DATA_BLOCK "Library: Part Numbers as Text"   // DB3
{ S7_Optimized_Access := 'TRUE' }
VERSION : 0.1
BEGIN
   pnText[0] := WSTRING#'';
   pnText[1] := WSTRING#'11.52.001.0545.000B';
   pnText[2] := WSTRING#'11.52.001.315.000B';
   pnText[3] := WSTRING#'11.52.001.316.001D';
   pnText[4] := WSTRING#'11.54.007.045.015D';
   pnText[5] := WSTRING#'11.54.007.052.007B';
   pnText[6] := WSTRING#'11.54.007.052.008A';
   pnText[7] := WSTRING#'11.54.007.052.009B';
   pnText[8] := WSTRING#'11.54.007.052.010B';
   pnText[9] := WSTRING#'11.54.007.315.026G';
   pnText[10] := WSTRING#'11.54.017.315.001F';
   pnText[11] := WSTRING#'16.08.208.011.010G';
   pnText[12] := WSTRING#'16.08.208.021.020C';
   pnText[13] := WSTRING#'16.08.208.031.020C';
   pnText[14] := WSTRING#'16.08.208.041.000A';
   pnText[15] := WSTRING#'16.08.208.051.000A';
   pnText[16] := WSTRING#'16.08.208.081.010B';
   pnText[17] := WSTRING#'16.08.208.091.000A';
   pnText[18] := WSTRING#'16.08.208.101.010C';
   pnText[19] := WSTRING#'16.08.208.111.000B';
   pnText[20] := WSTRING#'16.08.208.131.010L';
   pnText[21] := WSTRING#'16.08.208.151.010F';
   pnText[22] := WSTRING#'16.08.208.161.020F';
   pnText[23] := WSTRING#'16.08.208.301.000F';
   pnText[24] := WSTRING#'16.08.208.311.000F';
   pnText[25] := WSTRING#'16.08.208.321.000G';
   pnText[26] := WSTRING#'16.08.208.331.000F';
   pnText[27] := WSTRING#'16.08.208.411.030C';
   pnText[28] := WSTRING#'16.08.208.501.000B';
   pnText[29] := WSTRING#'16.08.208.531.020L';
   pnText[30] := WSTRING#'16.08.208.621.010C';
   pnText[31] := WSTRING#'16.08.208.631.000F';
   pnText[32] := WSTRING#'16.08.208.651.010B';
   pnText[33] := WSTRING#'16.08.208.661.000F';
   pnText[34] := WSTRING#'16.08.208.691.010D';
   pnText[35] := WSTRING#'16.08.209.031.010C';
   pnText[36] := WSTRING#'16.08.209.031.030B';
   pnText[37] := WSTRING#'16.08.209.031.050A';
   pnText[38] := WSTRING#'16.08.209.091.010C';
   pnText[39] := WSTRING#'16.08.209.091.030D';
   pnText[40] := WSTRING#'16.08.209.091.060A';
   pnText[41] := WSTRING#'16.08.209.232.010C';
   pnText[42] := WSTRING#'16.08.210.031.010B';
   pnText[43] := WSTRING#'16.08.210.421.010A';
   pnText[44] := WSTRING#'16.08.210.421.020A';
   pnText[45] := WSTRING#'16.08.210.421.030A';
   pnText[46] := WSTRING#'16.08.211.121.000G';
   pnText[47] := WSTRING#'16.08.211.291.000A';
   pnText[48] := WSTRING#'16.08.211.511.020F';
   pnText[49] := WSTRING#'16.08.211.551.000B';
   pnText[50] := WSTRING#'16.08.211.781.000A';
   pnText[51] := WSTRING#'16.08.211.801.010A';
   pnText[52] := WSTRING#'16.08.211.801.020A';
   pnText[53] := WSTRING#'16.08.211.806.020A';
   pnText[54] := WSTRING#'16.08.215.141.010C';
   pnText[55] := WSTRING#'16.08.215.871.010C';
   pnText[56] := WSTRING#'16.08.216.011.030B';
   pnText[57] := WSTRING#'16.08.216.053.000A';
   pnText[58] := WSTRING#'16.08.216.057.001A';
   pnText[59] := WSTRING#'16.08.216.141.010C';
   pnText[60] := WSTRING#'16.08.216.151.010B';
   pnText[61] := WSTRING#'16.08.216.161.020A';
   pnText[62] := WSTRING#'16.08.216.181.010B';
   pnText[63] := WSTRING#'16.08.216.181.090A';
   pnText[64] := WSTRING#'16.08.216.181.100A';
   pnText[65] := WSTRING#'16.08.216.181.110B';
   pnText[66] := WSTRING#'16.08.216.200.050A';
   pnText[67] := WSTRING#'16.08.216.202.080A';
   pnText[68] := WSTRING#'16.08.216.231.000B';
   pnText[69] := WSTRING#'16.08.216.251.000B';
   pnText[70] := WSTRING#'16.08.216.291.000A';
   pnText[71] := WSTRING#'16.08.216.315.000A';
   pnText[72] := WSTRING#'16.08.216.315.001A';
   pnText[73] := WSTRING#'16.08.216.315.002A';
   pnText[74] := WSTRING#'16.08.216.501.000C';
   pnText[75] := WSTRING#'16.08.216.501.010A';
   pnText[76] := WSTRING#'16.08.216.511.000C';
   pnText[77] := WSTRING#'16.08.216.515.008C';
   pnText[78] := WSTRING#'16.08.216.521.000C';
   pnText[79] := WSTRING#'16.08.216.526.002C';
   pnText[80] := WSTRING#'16.08.216.526.009A';
   pnText[81] := WSTRING#'16.08.216.551.000B';
   pnText[82] := WSTRING#'16.08.216.722.001A';
   pnText[83] := WSTRING#'16.08.216.790.001A';
   pnText[84] := WSTRING#'16.08.216.806.020A';
   pnText[85] := WSTRING#'16.08.216.831.020A';
   pnText[86] := WSTRING#'16.08.216.871.010C';
   pnText[87] := WSTRING#'16.08.216.910.020B';
   pnText[88] := WSTRING#'16.08.216.911.000C';
   pnText[89] := WSTRING#'16.08.216.911.000G';
   pnText[90] := WSTRING#'16.08.216.911.000H';
   pnText[91] := WSTRING#'16.08.216.911.030B';
   pnText[92] := WSTRING#'16.08.216.911.040B';
   pnText[93] := WSTRING#'16.08.216.912.050A';
   pnText[94] := WSTRING#'16.08.216.912.060B';
   pnText[95] := WSTRING#'16.08.216.951.010A';
   pnText[96] := WSTRING#'16.08.216.181.020A';
   pnText[97] := WSTRING#'16.08.217.411.080A';
   pnText[98] := WSTRING#'16.08.217.421.010A';
   pnText[99] := WSTRING#'16.08.217.421.130A';
   pnText[100] := WSTRING#'16.18.007.301.010A';
   pnText[101] := WSTRING#'16.18.007.301.020A';
   pnText[102] := WSTRING#'16.18.007.311.010A';
   pnText[103] := WSTRING#'16.18.007.311.020A';
   pnText[104] := WSTRING#'16.18.007.321.010B';
   pnText[105] := WSTRING#'16.18.008.301.010A';
   pnText[106] := WSTRING#'16.18.008.301.020A';
   pnText[107] := WSTRING#'16.18.008.301.030A';
   pnText[108] := WSTRING#'16.18.008.311.010A';
   pnText[109] := WSTRING#'16.18.008.311.020B';
   pnText[110] := WSTRING#'16.18.009.301.010A';
   pnText[111] := WSTRING#'16.18.009.301.020B';
   pnText[112] := WSTRING#'16.18.009.301.030A';
   pnText[113] := WSTRING#'16.18.009.301.040B';
   pnText[114] := WSTRING#'16.18.009.301.050A';
   pnText[115] := WSTRING#'16.18.009.311.010A';
   pnText[116] := WSTRING#'16.18.009.321.010A';
   pnText[117] := WSTRING#'16.18.009.321.020B';
   pnText[118] := WSTRING#'16.18.009.321.030A';
   pnText[119] := WSTRING#'16.18.009.331.030A';
   pnText[120] := WSTRING#'16.18.009.331.050A';
   pnText[121] := WSTRING#'16.18.009.371.010A';
   pnText[122] := WSTRING#'16.18.011.301.010A';
   pnText[123] := WSTRING#'16.18.011.301.020B';
   pnText[124] := WSTRING#'16.18.011.301.030A';
   pnText[125] := WSTRING#'16.18.011.301.040B';
   pnText[126] := WSTRING#'16.18.011.311.020A';
   pnText[127] := WSTRING#'16.18.011.321.010A';
   pnText[128] := WSTRING#'16.18.011.321.020B';
   pnText[129] := WSTRING#'16.18.011.321.030A';
   pnText[130] := WSTRING#'16.18.011.331.010A';
   pnText[131] := WSTRING#'16.18.011.331.020D';
   pnText[132] := WSTRING#'16.18.012.401.010A';
   pnText[133] := WSTRING#'16.18.012.401.020A';
   pnText[134] := WSTRING#'16.18.012.411.010A';
   pnText[135] := WSTRING#'16.18.012.411.020B';
   pnText[136] := WSTRING#'16.18.012.431.010A';
   pnText[137] := WSTRING#'16.18.012.441.010A';
   pnText[138] := WSTRING#'16.18.013.411.010A';
   pnText[139] := WSTRING#'16.18.013.411.020B';
   pnText[140] := WSTRING#'16.18.013.411.030A';
   pnText[141] := WSTRING#'16.18.013.421.010A';
   pnText[142] := WSTRING#'16.18.014.411.010A';
   pnText[143] := WSTRING#'16.18.014.411.030A';
   pnText[144] := WSTRING#'16.18.015.401.010A';
   pnText[145] := WSTRING#'16.18.015.411.010A';
   pnText[146] := WSTRING#'16.18.015.411.020B';
   pnText[147] := WSTRING#'16.18.015.411.030A';
   pnText[148] := WSTRING#'16.18.015.421.010A';
   pnText[149] := WSTRING#'16.18.015.421.020B';
   pnText[150] := WSTRING#'16.18.017.301.010A';
   pnText[151] := WSTRING#'16.18.017.301.020A';
   pnText[152] := WSTRING#'16.18.017.301.030A';
   pnText[153] := WSTRING#'16.18.017.301.040A';
   pnText[154] := WSTRING#'16.18.017.301.050A';
   pnText[155] := WSTRING#'16.18.017.311.010A';
   pnText[156] := WSTRING#'16.18.017.321.010A';
   pnText[157] := WSTRING#'16.18.017.321.020A';
   pnText[158] := WSTRING#'16.18.018.400.000A';
   pnText[159] := WSTRING#'16.18.018.401.010A';
   pnText[160] := WSTRING#'16.18.018.401.020B';
   pnText[161] := WSTRING#'16.18.018.401.030A';
   pnText[162] := WSTRING#'16.18.018.411.010A';
   pnText[163] := WSTRING#'16.18.018.421.010B';
   pnText[164] := WSTRING#'16.32.112.054.041A';
   pnText[165] := WSTRING#'16.32.112.057.010A';
   pnText[166] := WSTRING#'16.32.112.500.060D';
   pnText[167] := WSTRING#'16.32.112.500.090B';
   pnText[168] := WSTRING#'16.32.112.500.100A';
   pnText[169] := WSTRING#'16.32.112.500.120A';
   pnText[170] := WSTRING#'16.32.112.500.150B';
   pnText[171] := WSTRING#'16.32.112.500.160A';
   pnText[172] := WSTRING#'16.32.112.500.220A';
   pnText[173] := WSTRING#'16.32.112.500.300E';
   pnText[174] := WSTRING#'16.32.112.500.520B';
   pnText[175] := WSTRING#'16.32.112.502.050B';
   pnText[176] := WSTRING#'16.32.112.502.060B';
   pnText[177] := WSTRING#'16.32.112.502.070E';
   pnText[178] := WSTRING#'16.32.112.503.210A';
   pnText[179] := WSTRING#'16.32.112.503.220A';
   pnText[180] := WSTRING#'16.32.112.504.060A';
   pnText[181] := WSTRING#'16.32.112.504.070G';
   pnText[182] := WSTRING#'16.32.112.509.050E';
   pnText[183] := WSTRING#'16.32.112.509.070A';
   pnText[184] := WSTRING#'16.32.112.509.080F';
   pnText[185] := WSTRING#'16.32.112.516.110E';
   pnText[186] := WSTRING#'16.32.112.520.300E';
   pnText[187] := WSTRING#'16.32.112.521.010B';
   pnText[188] := WSTRING#'16.32.112.521.020B';
   pnText[189] := WSTRING#'16.32.112.521.030A';
   pnText[190] := WSTRING#'16.32.112.522.040D';
   pnText[191] := WSTRING#'16.32.112.522.050A';
   pnText[192] := WSTRING#'16.32.112.522.130A';
   pnText[193] := WSTRING#'16.32.112.529.010A';
   pnText[194] := WSTRING#'16.32.112.529.020B';
   pnText[195] := WSTRING#'16.32.112.529.030A';
   pnText[196] := WSTRING#'16.32.112.529.050D';
   pnText[197] := WSTRING#'16.32.112.536.010A';
   pnText[198] := WSTRING#'16.32.112.543.020A';
   pnText[199] := WSTRING#'16.32.112.543.210E';
   pnText[200] := WSTRING#'16.32.112.553.010A';
   pnText[201] := WSTRING#'16.32.112.553.020A';
   pnText[202] := WSTRING#'16.32.112.553.100D';
   pnText[203] := WSTRING#'16.32.112.553.220A';
   pnText[204] := WSTRING#'16.32.112.580.020A';
   pnText[205] := WSTRING#'16.32.112.601.030A';
   pnText[206] := WSTRING#'16.32.112.601.040A';
   pnText[207] := WSTRING#'16.32.112.621.010A';
   pnText[208] := WSTRING#'16.32.112.621.020A';
   pnText[209] := WSTRING#'16.32.112.704.000C';
   pnText[210] := WSTRING#'16.32.112.751.000D';
   pnText[211] := WSTRING#'16.32.112.751.001C';
   pnText[212] := WSTRING#'16.32.112.757.000A';
   pnText[213] := WSTRING#'16.32.112.757.001A';
   pnText[214] := WSTRING#'16.32.112.851.000A';
   pnText[215] := WSTRING#'16.32.112.851.001A';
   pnText[216] := WSTRING#'16.32.112.870.000C';
   pnText[217] := WSTRING#'16.32.307.211.150B';
   pnText[218] := WSTRING#'16.32.307.211.170B';
   pnText[219] := WSTRING#'16.32.307.212.320C';
   pnText[220] := WSTRING#'16.32.307.232.300B';
   pnText[221] := WSTRING#'16.32.307.262.300B';
   pnText[222] := WSTRING#'16.32.307.312.310A';
   pnText[223] := WSTRING#'16.32.307.461.160A';
   pnText[224] := WSTRING#'16.32.407.241.150B';
   pnText[225] := WSTRING#'16.32.407.241.170B';
   pnText[226] := WSTRING#'16.32.407.441.160A';
   pnText[227] := WSTRING#'16.32.606.311.010C';
   pnText[228] := WSTRING#'16.32.606.311.040B';
   pnText[229] := WSTRING#'16.32.606.311.050B';
   pnText[230] := WSTRING#'16.32.606.311.060A';
   pnText[231] := WSTRING#'16.32.606.311.070A';
   pnText[232] := WSTRING#'16.32.606.321.010B';
   pnText[233] := WSTRING#'16.32.606.321.030B';
   pnText[234] := WSTRING#'16.32.706.311.010C';
   pnText[235] := WSTRING#'16.32.706.311.020B';
   pnText[236] := WSTRING#'16.32.706.311.040B';
   pnText[237] := WSTRING#'16.32.706.311.050B';
   pnText[238] := WSTRING#'16.32.706.321.010B';
   pnText[239] := WSTRING#'16.32.706.321.030B';
   pnText[240] := WSTRING#'16.32.706.401.040A';
   pnText[241] := WSTRING#'16.32.706.401.050A';
   pnText[242] := WSTRING#'16.32.806.502.080A';
   pnText[243] := WSTRING#'DUNNAGE';
   pnText[244] := WSTRING#'PEANUTS';
   pnText[245] := WSTRING#'RINGS CART';
END_DATA_BLOCK

DATA_BLOCK "LED Sign"   // DB4
{ S7_Optimized_Access := 'TRUE' }
VERSION : 0.1
   VAR
      request : "LED Sign Data";
   END_VAR
BEGIN
END_DATA_BLOCK

DATA_BLOCK "HMI Stations: Saved Wips"   // DB5
{ S7_Optimized_Access := 'TRUE' }
VERSION : 0.1
BEGIN
   stn[0].pStn := 25;
   stn[1].pStn := 26;
   stn[2].pStn := 27;
   stn[3].pStn := 28;
   stn[4].pStn := 29;
END_DATA_BLOCK

DATA_BLOCK "HMI Data: TP700 Stations"   // DB6
{ S7_Optimized_Access := 'TRUE' }
VERSION : 0.1
BEGIN
END_DATA_BLOCK

DATA_BLOCK "Library: Wip Names as Text"   // DB8
{ S7_Optimized_Access := 'TRUE' }
VERSION : 0.1
BEGIN
   code[0] := WSTRING#'';
   code[1] := WSTRING#'11.52.001.312.000B';
   code[2] := WSTRING#'11.54.007.309.000D';
   code[3] := WSTRING#'11.54.007.309.002D';
   code[4] := WSTRING#'16.08.208.031.000F';
   code[5] := WSTRING#'16.08.208.081.000H';
   code[6] := WSTRING#'16.08.208.101.020A';
   code[7] := WSTRING#'16.08.208.621.000G';
   code[8] := WSTRING#'16.08.208.651.000G';
   code[9] := WSTRING#'16.08.209.031.000C';
   code[10] := WSTRING#'16.08.209.091.000D';
   code[11] := WSTRING#'16.08.209.233.000E';
   code[12] := WSTRING#'16.08.209.437.000A';
   code[13] := WSTRING#'16.08.210.031.000B';
   code[14] := WSTRING#'16.08.210.421.500A';
   code[15] := WSTRING#'16.08.210.428.000A';
   code[16] := WSTRING#'16.08.211.801.400A';
   code[17] := WSTRING#'16.08.211.801.700B';
   code[18] := WSTRING#'16.08.211.803.400A';
   code[19] := WSTRING#'16.08.211.806.400B';
   code[20] := WSTRING#'16.08.216.751.100A';
   code[21] := WSTRING#'16.08.216.801.600A';
   code[22] := WSTRING#'16.08.216.806.400A';
   code[23] := WSTRING#'16.08.217.233.000A';
   code[24] := WSTRING#'16.08.217.408.000A';
   code[25] := WSTRING#'16.08.217.421.500A';
   code[26] := WSTRING#'16.08.217.737.000A';
   code[27] := WSTRING#'16.18.007.300.000A';
   code[28] := WSTRING#'16.18.007.310.000A';
   code[29] := WSTRING#'16.18.007.320.000B';
   code[30] := WSTRING#'16.18.008.300.000A';
   code[31] := WSTRING#'16.18.008.310.000A';
   code[32] := WSTRING#'16.18.008.320.000A';
   code[33] := WSTRING#'16.18.008.340.000A';
   code[34] := WSTRING#'16.18.009.301.000H';
   code[35] := WSTRING#'16.18.009.311.000H';
   code[36] := WSTRING#'16.18.009.321.000G';
   code[37] := WSTRING#'16.18.009.331.000F';
   code[38] := WSTRING#'16.18.009.371.000D';
   code[39] := WSTRING#'16.18.011.300.000A';
   code[40] := WSTRING#'16.18.011.310.000A';
   code[41] := WSTRING#'16.18.011.320.000A';
   code[42] := WSTRING#'16.18.011.330.000A';
   code[43] := WSTRING#'16.18.011.340.000A';
   code[44] := WSTRING#'16.18.012.400.000A';
   code[45] := WSTRING#'16.18.012.410.000A';
   code[46] := WSTRING#'16.18.012.420.000A';
   code[47] := WSTRING#'16.18.012.430.000A';
   code[48] := WSTRING#'16.18.012.440.000A';
   code[49] := WSTRING#'16.18.013.410.000A';
   code[50] := WSTRING#'16.18.013.420.000A';
   code[51] := WSTRING#'16.18.015.400.000A';
   code[52] := WSTRING#'16.18.015.410.000A';
   code[53] := WSTRING#'16.18.015.420.000A';
   code[54] := WSTRING#'16.18.015.430.000A';
   code[55] := WSTRING#'16.18.015.450.000A';
   code[56] := WSTRING#'16.18.016.400.000A';
   code[57] := WSTRING#'16.18.017.300.000A';
   code[58] := WSTRING#'16.18.017.310.000A';
   code[59] := WSTRING#'16.18.017.321.000F';
   code[60] := WSTRING#'16.18.018.400.000A';
   code[61] := WSTRING#'16.18.018.410.000A';
   code[62] := WSTRING#'16.18.018.420.000A';
   code[63] := WSTRING#'16.18.018.440.000A';
   code[64] := WSTRING#'16.32.112.304.008A';
   code[65] := WSTRING#'16.32.112.311.001A';
   code[66] := WSTRING#'16.32.112.516.000G';
   code[67] := WSTRING#'16.32.112.543.000E';
   code[68] := WSTRING#'16.32.112.553.300C';
   code[69] := WSTRING#'16.32.307.322.210A';
   code[70] := WSTRING#'16.32.307.332.300A';
   code[71] := WSTRING#'16.32.307.332.400A';
   code[72] := WSTRING#'16.32.307.472.210A';
   code[73] := WSTRING#'16.32.407.322.210A';
   code[74] := WSTRING#'16.32.407.322.300A';
   code[75] := WSTRING#'16.32.606.411.000A';
   code[76] := WSTRING#'16.32.606.421.000A';
   code[77] := WSTRING#'16.32.706.311.000A';
   code[78] := WSTRING#'16.32.706.311.001A';
   code[79] := WSTRING#'16.32.706.341.000A';
   code[80] := WSTRING#'16.32.706.401.000A';
   txt[0] := WSTRING#'NO TEXT ENTERED';
   txt[1] := WSTRING#'DPF Sleeved 2016';
   txt[2] := WSTRING#'SA SCR CANNING 9.5 x 10in -END FORMED-';
   txt[3] := WSTRING#'Assembly DPF Canning 2016';
   txt[4] := WSTRING#'ASSY DOC CANNING A700';
   txt[5] := WSTRING#'ASSY DPF CANNING A700';
   txt[6] := WSTRING#'ASSY SCR CANNING FORMED';
   txt[7] := WSTRING#'DOC Stuffed Shell Before Forming';
   txt[8] := WSTRING#'DOC Stuffed Shell Unformed';
   txt[9] := WSTRING#'DPF Stuffed Shell 1 box longs only';
   txt[10] := WSTRING#'DPF Stuffed Shell MD11';
   txt[11] := WSTRING#'DPF Stuffed Shell: MD13/MD16';
   txt[12] := WSTRING#'SA DOC CANNING 11.25 x 3.4in -END FORMED';
   txt[13] := WSTRING#'SA DOC CANNING 11.25 x 4in -END FORMED-';
   txt[14] := WSTRING#'SA DOC CANNING 11.25 x 5in -END FORMED-';
   txt[15] := WSTRING#'SA DOC CANNING 11.25 x 6.8in -END FORMED';
   txt[16] := WSTRING#'SA DOC CANNING 11_25 x 5in -END FORMED-';
   txt[17] := WSTRING#'SA DOC CANNING 9.5 x 3.3in -END FORMED-';
   txt[18] := WSTRING#'SA DOC CANNING 9.5 x 4in -END FORMED-';
   txt[19] := WSTRING#'SA DOC CANNING 9.5 x 4in -END FORMED_';
   txt[20] := WSTRING#'SA DOC CANNING 9.5 x 5.5in -END FORMED-';
   txt[21] := WSTRING#'SA DOC CANNING 9.5 x 5in -END FORMED-';
   txt[22] := WSTRING#'SA DOC CANNING 9_5 x 4_5in -END FORMED-';
   txt[23] := WSTRING#'SA DOC Canning w/out End Forming';
   txt[24] := WSTRING#'SA DOC Sleeved';
   txt[25] := WSTRING#'SA DOC SLEEVED - 2HH 2016';
   txt[26] := WSTRING#'SA DOC SLEEVED - 2V2 2016 unformed';
   txt[27] := WSTRING#'SA DOC Sleeved Before Forming';
   txt[28] := WSTRING#'SA DOC Sleeved DDC 2016 unformed';
   txt[29] := WSTRING#'SA DPF SLEEVED Hess';
   txt[30] := WSTRING#'SA DPF Stuffed (after Hess)';
   txt[31] := WSTRING#'SA DPF Stuffed Shell';
   txt[32] := WSTRING#'SA JL 2.2L DPF CANNING';
   txt[33] := WSTRING#'SA SCR CANNING 12 x 10in -END FORMED-';
   txt[34] := WSTRING#'SA SCR CANNING 12 x 9in -END FORMED-';
   txt[35] := WSTRING#'SA SCR CANNING 12x7in UNFORMED-';
   txt[36] := WSTRING#'SA SCR CANNING 13 x 11in UNFORMED-';
   txt[37] := WSTRING#'SA SCR CANNING 13 x 12in UNFORMED-';
   txt[38] := WSTRING#'SA SCR CANNING 13 x 9in UNFORMED';
   txt[39] := WSTRING#'SA SCR CANNING 13 X10 UNFORMED';
   txt[40] := WSTRING#'SA SCR CANNING 9.5 x 10in -END FORMED-';
   txt[41] := WSTRING#'SA SCR CANNING 9.5 x 12in -END FORMED-';
   txt[42] := WSTRING#'SA SCR CANNING 9.5 x 13.5in -END FORMED-';
   txt[43] := WSTRING#'SA SCR CANNING 9.5 x 13in -END FORMED-';
   txt[44] := WSTRING#'SA SCR CANNING 9.5 x 9in -END FORMED-';
   txt[45] := WSTRING#'SA SCR CANNING 9_5 x 13in -END FORMED-';
   txt[46] := WSTRING#'SA SCR CANNING A700 UNFORMED';
   txt[47] := WSTRING#'SA SCR CANNING UNFORMED';
   txt[48] := WSTRING#'SA SCR Catalyst Module - MD11_MD13 -';
   txt[49] := WSTRING#'SA SCR SLEEVED before FORMING';
   txt[50] := WSTRING#'SA Sleeved SCR 2016';
   txt[51] := WSTRING#'SCR CANNING 9.5 x 9in -END FORMED-';
   txt[52] := WSTRING#'SCR Stuffed Shell 1 box longs only';
   txt[53] := WSTRING#'SCR Stuffed Shell High Power';
   txt[54] := WSTRING#'SCR Stuffed Shell MD11/13: Australia';
   txt[55] := WSTRING#'SCR Stuffed Shell MD11/13: Vert Short';
   txt[56] := WSTRING#'SCR Stuffed Shell- NGK Before Forming';
   txt[57] := WSTRING#'Stuffed Shell - SCR Horizontal';
   txt[58] := WSTRING#'Stuffed Shell - SCR Horizontal Long- UNI';
   txt[59] := WSTRING#'STUFFED SHELL ASSEMBLY USA-U625';
   txt[60] := WSTRING#'Stuffed Shell DOC';
   txt[61] := WSTRING#'Stuffed Shell DOC- 2013';
   txt[62] := WSTRING#'Stuffed Shell SCR- NGK';
   txt[63] := WSTRING#'Volvo - ASSY INLET - SUB 8 Unformed';
   txt[64] := WSTRING#'VOLVO DOC STUFFED SHELL UNFORMED';
END_DATA_BLOCK

DATA_BLOCK "Stations"   // DB10
{ S7_Optimized_Access := 'TRUE' }
VERSION : 0.1
BEGIN
   stn[0].id.dropZone := 1;
   stn[0].id.lineName := WSTRING#'VOLVO 16';
   stn[1].id.dropZone := 2;
   stn[1].id.lineName := WSTRING#'VOLVO 16';
   stn[2].id.dropZone := 3;
   stn[2].id.lineName := WSTRING#'VOLVO 16';
   stn[3].id.dropZone := 4;
   stn[3].id.lineName := WSTRING#'VOLVO 16';
   stn[4].id.dropZone := 5;
   stn[4].id.lineName := WSTRING#'VOLVO 16';
   stn[5].id.dropZone := 6;
   stn[5].id.lineName := WSTRING#'VOLVO 16';
   stn[6].id.dropZone := 7;
   stn[6].id.lineName := WSTRING#'VOLVO 16';
   stn[7].id.dropZone := 8;
   stn[7].id.lineName := WSTRING#'VOLVO 16';
   stn[8].id.dropZone := 9;
   stn[8].id.lineName := WSTRING#'VOLVO 16';
   stn[9].id.dropZone := 10;
   stn[9].id.lineName := WSTRING#'VOLVO 16';
   stn[10].id.dropZone := 11;
   stn[10].id.lineName := WSTRING#'VOLVO 16';
   stn[11].id.dropZone := 1;
   stn[11].id.lineName := WSTRING#'CHM';
   stn[12].id.dropZone := 2;
   stn[12].id.lineName := WSTRING#'CHM';
   stn[13].id.dropZone := 3;
   stn[13].id.lineName := WSTRING#'CHM';
   stn[14].id.dropZone := 4;
   stn[14].id.lineName := WSTRING#'CHM';
   stn[15].id.dropZone := 5;
   stn[15].id.lineName := WSTRING#'CHM';
   stn[16].id.dropZone := 1;
   stn[16].id.lineName := WSTRING#'CDO';
   stn[17].id.dropZone := 2;
   stn[17].id.lineName := WSTRING#'CDO';
   stn[18].id.dropZone := 3;
   stn[18].id.lineName := WSTRING#'CDO';
   stn[19].id.dropZone := 1;
   stn[19].id.lineName := WSTRING#'BFL';
   stn[20].id.dropZone := 2;
   stn[20].id.lineName := WSTRING#'BFL';
   stn[21].id.dropZone := 3;
   stn[21].id.lineName := WSTRING#'BFL';
   stn[22].id.dropZone := 1;
   stn[22].id.lineName := WSTRING#'LGS';
   stn[23].id.dropZone := 2;
   stn[23].id.lineName := WSTRING#'LGS';
   stn[24].id.dropZone := 3;
   stn[24].id.lineName := WSTRING#'LGS';
   stn[25].id.dropZone := 1;
   stn[25].id.lineName := WSTRING#'CV';
   stn[25].wipData.index := -1;
   stn[26].id.dropZone := 2;
   stn[26].id.lineName := WSTRING#'CV';
   stn[27].id.dropZone := 3;
   stn[27].id.lineName := WSTRING#'CV';
   stn[28].id.dropZone := 4;
   stn[28].id.lineName := WSTRING#'CV';
   stn[29].id.dropZone := 1;
   stn[29].id.lineName := WSTRING#'PC';
   stn[30].id.dropZone := 2;
   stn[30].id.lineName := WSTRING#'PC';
   stn[31].id.dropZone := 1;
   stn[31].id.lineName := WSTRING#'1BX2.0';
   stn[32].id.dropZone := 2;
   stn[32].id.lineName := WSTRING#'1BX2.0';
   stn[33].id.dropZone := 3;
   stn[33].id.lineName := WSTRING#'1BX2.0';
   stn[34].id.dropZone := 4;
   stn[34].id.lineName := WSTRING#'1BX2.0';
   stn[35].id.dropZone := 5;
   stn[35].id.lineName := WSTRING#'1BX2.0';
   stn[36].id.dropZone := 1;
   stn[36].id.lineName := WSTRING#'1BX3.0';
   stn[37].id.dropZone := 2;
   stn[37].id.lineName := WSTRING#'1BX3.0';
   stn[38].id.lineName := WSTRING#'1BX3.0';
   stn[38].id.dropZone := 3;
END_DATA_BLOCK

DATA_BLOCK "Part Requests"   // DB11
{ S7_Optimized_Access := 'TRUE' }
VERSION : 0.1
BEGIN
   row[0] := -1;
   row[1] := -1;
   row[2] := -1;
   row[3] := -1;
   row[4] := -1;
   row[5] := -1;
   row[6] := -1;
   row[7] := -1;
   row[8] := -1;
   row[9] := -1;
   row[10] := -1;
   row[11] := -1;
   row[12] := -1;
   row[13] := -1;
   row[14] := -1;
   row[15] := -1;
   row[16] := -1;
   row[17] := -1;
   row[18] := -1;
   row[19] := -1;
   row[20] := -1;
   row[21] := -1;
   row[22] := -1;
   row[23] := -1;
   row[24] := -1;
   row[25] := -1;
   row[26] := -1;
   row[27] := -1;
   row[28] := -1;
   row[29] := -1;
   row[30] := -1;
   row[31] := -1;
   row[32] := -1;
   row[33] := -1;
   row[34] := -1;
   row[35] := -1;
   row[36] := -1;
   row[37] := -1;
   row[38] := -1;
   row[39] := -1;
   row[40] := -1;
   row[41] := -1;
   row[42] := -1;
   row[43] := -1;
   row[44] := -1;
   row[45] := -1;
   row[46] := -1;
   row[47] := -1;
   row[48] := -1;
   row[49] := -1;
   row[50] := -1;
   row[51] := -1;
   row[52] := -1;
   row[53] := -1;
   row[54] := -1;
   row[55] := -1;
   row[56] := -1;
   row[57] := -1;
   row[58] := -1;
   row[59] := -1;
   row[60] := -1;
   row[61] := -1;
   row[62] := -1;
   row[63] := -1;
   row[64] := -1;
   row[65] := -1;
   row[66] := -1;
   row[67] := -1;
   row[68] := -1;
   row[69] := -1;
   row[70] := -1;
   row[71] := -1;
   row[72] := -1;
   row[73] := -1;
   row[74] := -1;
   row[75] := -1;
   row[76] := -1;
   row[77] := -1;
   row[78] := -1;
   row[79] := -1;
   row[80] := -1;
   row[81] := -1;
   row[82] := -1;
   row[83] := -1;
   row[84] := -1;
   row[85] := -1;
   row[86] := -1;
   row[87] := -1;
   row[88] := -1;
   row[89] := -1;
   row[90] := -1;
   row[91] := -1;
   row[92] := -1;
   row[93] := -1;
   row[94] := -1;
   row[95] := -1;
   row[96] := -1;
   row[97] := -1;
   row[98] := -1;
   row[99] := -1;
   row[100] := -1;
   row[101] := -1;
   row[102] := -1;
   row[103] := -1;
   row[104] := -1;
   row[105] := -1;
   row[106] := -1;
   row[107] := -1;
   row[108] := -1;
   row[109] := -1;
   row[110] := -1;
   row[111] := -1;
   row[112] := -1;
   row[113] := -1;
   row[114] := -1;
   row[115] := -1;
   row[116] := -1;
   row[117] := -1;
   row[118] := -1;
   row[119] := -1;
   row[120] := -1;
   row[121] := -1;
   row[122] := -1;
   row[123] := -1;
   row[124] := -1;
   row[125] := -1;
   row[126] := -1;
   row[127] := -1;
   row[128] := -1;
   row[129] := -1;
   row[130] := -1;
   row[131] := -1;
   row[132] := -1;
   row[133] := -1;
   row[134] := -1;
   row[135] := -1;
   row[136] := -1;
   row[137] := -1;
   row[138] := -1;
   row[139] := -1;
   row[140] := -1;
   row[141] := -1;
   row[142] := -1;
   row[143] := -1;
   row[144] := -1;
   row[145] := -1;
   row[146] := -1;
   row[147] := -1;
   row[148] := -1;
   row[149] := -1;
   row[150] := -1;
   row[151] := -1;
   row[152] := -1;
   row[153] := -1;
   row[154] := -1;
   row[155] := -1;
   row[156] := -1;
   row[157] := -1;
   row[158] := -1;
   row[159] := -1;
   row[160] := -1;
   row[161] := -1;
   row[162] := -1;
   row[163] := -1;
   row[164] := -1;
   row[165] := -1;
   row[166] := -1;
   row[167] := -1;
   row[168] := -1;
   row[169] := -1;
   row[170] := -1;
   row[171] := -1;
   row[172] := -1;
   row[173] := -1;
   row[174] := -1;
   row[175] := -1;
   row[176] := -1;
   row[177] := -1;
   row[178] := -1;
   row[179] := -1;
   row[180] := -1;
   row[181] := -1;
   row[182] := -1;
   row[183] := -1;
   row[184] := -1;
   row[185] := -1;
   row[186] := -1;
   row[187] := -1;
   row[188] := -1;
   row[189] := -1;
   row[190] := -1;
   row[191] := -1;
   row[192] := -1;
   row[193] := -1;
   row[194] := -1;
   row[195] := -1;
   row[196] := -1;
   row[197] := -1;
   row[198] := -1;
   row[199] := -1;
END_DATA_BLOCK

// folder: Test Area

DATA_BLOCK "Test DB"   // DB9
{ S7_Optimized_Access := 'TRUE' }
VERSION : 0.1
   VAR
      run_collapse_test : Bool;
      test_collapse_array : Array[0..9] of Int;
   END_VAR
BEGIN
   test_collapse_array[0] := 5;
   test_collapse_array[1] := -1;
   test_collapse_array[2] := 4;
   test_collapse_array[3] := -1;
   test_collapse_array[4] := -1;
   test_collapse_array[5] := -1;
   test_collapse_array[6] := -1;
   test_collapse_array[7] := -1;
   test_collapse_array[8] := 10;
   test_collapse_array[9] := 44;
END_DATA_BLOCK

// folder: (top level)

FUNCTION_BLOCK "EMP"   // FB1, LAD
{ S7_Optimized_Access := 'TRUE' }
VERSION : 0.1
   VAR
      "inst Global To Sim" : "Sim: from Global";
      "inst KP8 Button Activation" : "Button Parameters";
      "inst KP8 Drivers" : Array[0.."stnCount"] of "KP8 Driver";
      "inst Sim to Global" : "Sim: from Global";
      "inst Order States" : "Order State";
      "inst Flag Manager" : "Flag";
      "inst Order Timers" : "Order Timer";
      "inst HMI:Part Call: Table Driver" : "Part Call";
      "inst Part Request" : "Part Request";
      "inst HMI Station" : "HMI Station";
      "inst From Excel" : "From Excel";
      "Inst Settings Screen" : "Settings Screen";
      "inst Pop Up: Select Station_DB" : "Pop Up: Select Stations";
      "inst Pop Up: Select Buttons" : "Pop Up: Select Buttons";
      "inst Pop Up: Select WIPs" : "Pop Up: Select WIPs";
   END_VAR
   VAR_TEMP
      pStn : Int;
   END_VAR
BEGIN

REGION Network 1: SIMULATION TO GLOBAL
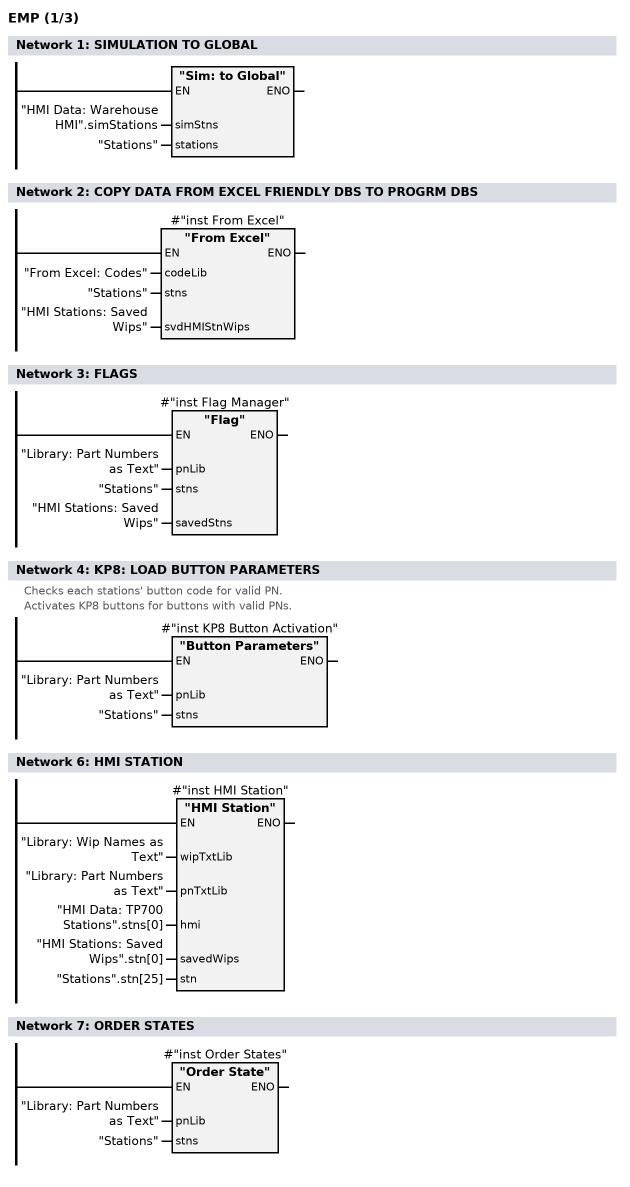
   RUNG wire#powerrail
      "Sim: to Global"(simStns := "HMI Data: Warehouse HMI".simStations, stations := "Stations")
   END_RUNG
   // the same network as SCL:
   "Sim: to Global"(simStns := "HMI Data: Warehouse HMI".simStations, stations := "Stations");
END_REGION

REGION Network 2: COPY DATA FROM EXCEL FRIENDLY DBS TO PROGRM DBS
   RUNG wire#powerrail
      #"inst From Excel"(codeLib := "From Excel: Codes", stns := "Stations", svdHMIStnWips := "HMI Stations: Saved Wips")
   END_RUNG
   // the same network as SCL:
   #"inst From Excel"(codeLib := "From Excel: Codes",   // "From Excel"
                      stns := "Stations",
                      svdHMIStnWips := "HMI Stations: Saved Wips");
END_REGION

REGION Network 3: FLAGS
   RUNG wire#powerrail
      #"inst Flag Manager"(pnLib := "Library: Part Numbers as Text", stns := "Stations", savedStns := "HMI Stations: Saved Wips")
   END_RUNG
   // the same network as SCL:
   #"inst Flag Manager"(pnLib := "Library: Part Numbers as Text",   // "Flag"
                        stns := "Stations",
                        savedStns := "HMI Stations: Saved Wips");
END_REGION

REGION Network 4: KP8: LOAD BUTTON PARAMETERS
   // Checks each stations' button code for valid PN.
   // Activates KP8 buttons for buttons with valid PNs.
   RUNG wire#powerrail
      #"inst KP8 Button Activation"(pnLib := "Library: Part Numbers as Text", stns := "Stations")
   END_RUNG
   // the same network as SCL:
   #"inst KP8 Button Activation"(pnLib := "Library: Part Numbers as Text", stns := "Stations");   // "Button Parameters"
END_REGION

REGION Network 5 (SCL): KP8 DRIVER CALLS
   // HMI stations do not use the KP8 driver and are skipped by the case statement.
   REGION "LOOP THROUGH STATIONS"
       FOR #pStn := 0 TO "stnCount" DO

           REGION "CALL ONLY FOR KP8 STATIONS"
               CASE #pStn OF
                   0..23,29.."stnCount":
                       #"inst KP8 Drivers"[#pStn](kp8DI := "Stations".stn[#pStn].wipCmpts.ioData.kp8.input,
                                                  "reset" := "Stations".stn[#pStn].wipCmpts.flags.resetStation,
                                                  btnParams := "Stations".stn[#pStn].kp8Config,
                                                  kp8DQ => "Stations".stn[#pStn].wipCmpts.ioData.kp8.tempOut,
                                                  physical => "Stations".stn[#pStn].kp8Physical,
                                                  logical => "Stations".stn[#pStn].wipCmpts.kp8Logical);
                   ELSE
                       ;
               END_CASE;
           END_REGION

       END_FOR;
   END_REGION
END_REGION

REGION Network 6: HMI STATION
   RUNG wire#powerrail
      #"inst HMI Station"(wipTxtLib := "Library: Wip Names as Text", pnTxtLib := "Library: Part Numbers as Text", hmi := "HMI Data: TP700 Stations".stns[0], savedWips := "HMI Stations: Saved Wips".stn[0], stn := "Stations".stn[25])
   END_RUNG
   // the same network as SCL:
   #"inst HMI Station"(wipTxtLib := "Library: Wip Names as Text",   // "HMI Station"
                       pnTxtLib := "Library: Part Numbers as Text",
                       hmi := "HMI Data: TP700 Stations".stns[0],
                       savedWips := "HMI Stations: Saved Wips".stn[0],
                       stn := "Stations".stn[25]);
END_REGION

REGION Network 7: ORDER STATES
   RUNG wire#powerrail
      #"inst Order States"(pnLib := "Library: Part Numbers as Text", stns := "Stations")
   END_RUNG
   // the same network as SCL:
   #"inst Order States"(pnLib := "Library: Part Numbers as Text", stns := "Stations");   // "Order State"
END_REGION

REGION Network 8: PART REQUESTS
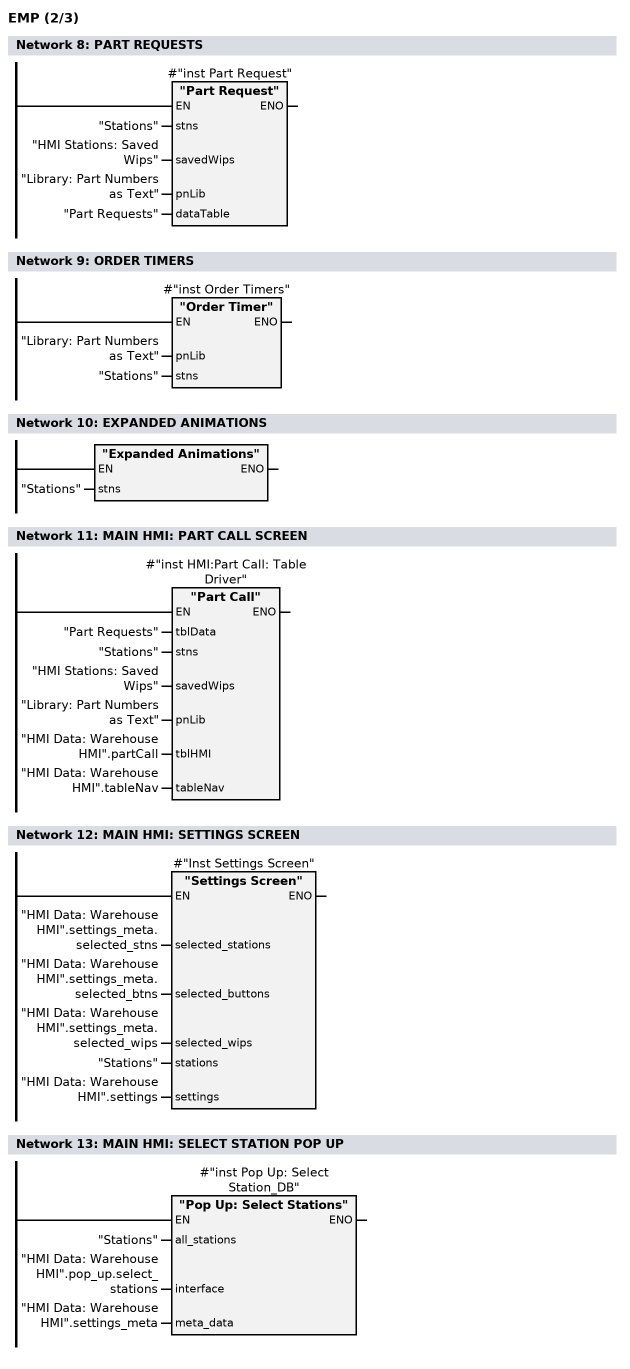
   RUNG wire#powerrail
      #"inst Part Request"(stns := "Stations", savedWips := "HMI Stations: Saved Wips", pnLib := "Library: Part Numbers as Text", dataTable := "Part Requests")
   END_RUNG
   // the same network as SCL:
   #"inst Part Request"(stns := "Stations",   // "Part Request"
                        savedWips := "HMI Stations: Saved Wips",
                        pnLib := "Library: Part Numbers as Text",
                        dataTable := "Part Requests");
END_REGION

REGION Network 9: ORDER TIMERS
   RUNG wire#powerrail
      #"inst Order Timers"(pnLib := "Library: Part Numbers as Text", stns := "Stations")
   END_RUNG
   // the same network as SCL:
   #"inst Order Timers"(pnLib := "Library: Part Numbers as Text", stns := "Stations");   // "Order Timer"
END_REGION

REGION Network 10: EXPANDED ANIMATIONS
   RUNG wire#powerrail
      "Expanded Animations"(stns := "Stations")
   END_RUNG
   // the same network as SCL:
   "Expanded Animations"(stns := "Stations");
END_REGION

REGION Network 11: MAIN HMI: PART CALL SCREEN
   RUNG wire#powerrail
      #"inst HMI:Part Call: Table Driver"(tblData := "Part Requests", stns := "Stations", savedWips := "HMI Stations: Saved Wips", pnLib := "Library: Part Numbers as Text", tblHMI := "HMI Data: Warehouse HMI".partCall, tableNav := "HMI Data: Warehouse HMI".tableNav)
   END_RUNG
   // the same network as SCL:
   #"inst HMI:Part Call: Table Driver"(tblData := "Part Requests",   // "Part Call"
                           stns := "Stations",
                           savedWips := "HMI Stations: Saved Wips",
                           pnLib := "Library: Part Numbers as Text",
                           tblHMI := "HMI Data: Warehouse HMI".partCall,
                           tableNav := "HMI Data: Warehouse HMI".tableNav);
END_REGION

REGION Network 12: MAIN HMI: SETTINGS SCREEN
   RUNG wire#powerrail
      #"Inst Settings Screen"(selected_stations := "HMI Data: Warehouse HMI".settings_meta.selected_stns, selected_buttons := "HMI Data: Warehouse HMI".settings_meta.selected_btns, selected_wips := "HMI Data: Warehouse HMI".settings_meta.selected_wips, stations := "Stations", settings := "HMI Data: Warehouse HMI".settings)
   END_RUNG
   // the same network as SCL:
   #"Inst Settings Screen"(selected_stations := "HMI Data: Warehouse HMI".settings_meta.selected_stns,   // "Settings Screen"
                           selected_buttons := "HMI Data: Warehouse HMI".settings_meta.selected_btns,
                           selected_wips := "HMI Data: Warehouse HMI".settings_meta.selected_wips,
                           stations := "Stations",
                           settings := "HMI Data: Warehouse HMI".settings);
END_REGION

REGION Network 13: MAIN HMI: SELECT STATION POP UP
   RUNG wire#powerrail
      #"inst Pop Up: Select Station_DB"(all_stations := "Stations", interface := "HMI Data: Warehouse HMI".pop_up.select_stations, meta_data := "HMI Data: Warehouse HMI".settings_meta)
   END_RUNG
   // the same network as SCL:
   #"inst Pop Up: Select Station_DB"(all_stations := "Stations",   // "Pop Up: Select Stations"
                           interface := "HMI Data: Warehouse HMI".pop_up.select_stations,
                           meta_data := "HMI Data: Warehouse HMI".settings_meta);
END_REGION

REGION Network 14: MAIN HMI: SELECT WIPS POP UP
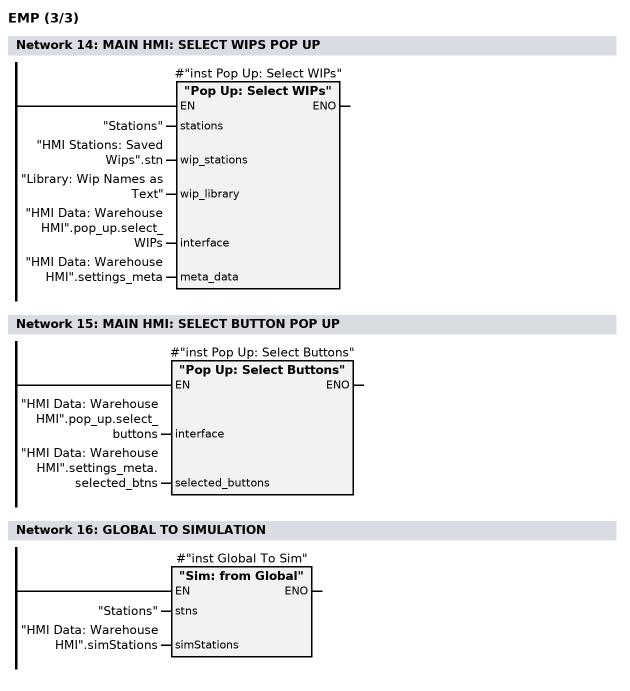
   RUNG wire#powerrail
      #"inst Pop Up: Select WIPs"(stations := "Stations", wip_stations := "HMI Stations: Saved Wips".stn, wip_library := "Library: Wip Names as Text", interface := "HMI Data: Warehouse HMI".pop_up.select_WIPs, meta_data := "HMI Data: Warehouse HMI".settings_meta)
   END_RUNG
   // the same network as SCL:
   #"inst Pop Up: Select WIPs"(stations := "Stations",   // "Pop Up: Select WIPs"
                           wip_stations := "HMI Stations: Saved Wips".stn,
                           wip_library := "Library: Wip Names as Text",
                           interface := "HMI Data: Warehouse HMI".pop_up.select_WIPs,
                           meta_data := "HMI Data: Warehouse HMI".settings_meta);
END_REGION

REGION Network 15: MAIN HMI: SELECT BUTTON POP UP
   RUNG wire#powerrail
      #"inst Pop Up: Select Buttons"(interface := "HMI Data: Warehouse HMI".pop_up.select_buttons, selected_buttons := "HMI Data: Warehouse HMI".settings_meta.selected_btns)
   END_RUNG
   // the same network as SCL:
   #"inst Pop Up: Select Buttons"(interface := "HMI Data: Warehouse HMI".pop_up.select_buttons,   // "Pop Up: Select Buttons"
                           selected_buttons := "HMI Data: Warehouse HMI".settings_meta.selected_btns);
END_REGION

REGION Network 16: GLOBAL TO SIMULATION
   RUNG wire#powerrail
      #"inst Global To Sim"(stns := "Stations", simStations := "HMI Data: Warehouse HMI".simStations)
   END_RUNG
   // the same network as SCL:
   #"inst Global To Sim"(stns := "Stations", simStations := "HMI Data: Warehouse HMI".simStations);   // "Sim: from Global"
END_REGION
END_FUNCTION_BLOCK

FUNCTION_BLOCK "Table"   // FB20, SCL
{ S7_Optimized_Access := 'TRUE' }
VERSION : 0.1
   VAR
      row_count : Int;
   END_VAR
BEGIN
END_FUNCTION_BLOCK

ORGANIZATION_BLOCK "Main"   // OB1, LAD, ProgramCycle
TITLE = "Main Program Sweep (Cycle)"
{ S7_Optimized_Access := 'TRUE' }
VERSION : 0.1
   VAR_INPUT
      Initial_Call : Bool;   // Initial call of this OB
      Remanence : Bool;   // =True, if remanent data are available
   END_VAR
BEGIN

REGION Network 1
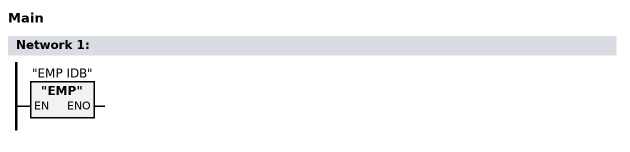
   RUNG wire#powerrail
      "EMP IDB"()
   END_RUNG
   // the same network as SCL:
   "EMP IDB"();   // "EMP"
END_REGION
END_ORGANIZATION_BLOCK

// folder: Flags

FUNCTION_BLOCK "Flag: New PN Code"   // FB3, SCL
{ S7_Optimized_Access := 'TRUE' }
VERSION : 0.1
   VAR_IN_OUT
      stns : "Station: All Stations";
   END_VAR
   VAR
      old : Struct
         pnCode : Array[0.."stnCount"] of Struct
            me : Array[0.."btnCount"] of DInt;
         END_STRUCT;
      END_STRUCT;
   END_VAR
   VAR_TEMP
      pStn : Int;
      ret : Bool;
   END_VAR
BEGIN
   REGION "FOR EACH STATION"
       FOR #pStn := 0 TO "stnCount" DO

           REGION "ON PART NUMBER CHANGE"
               IF #stns.stn[#pStn].wipCmpts.pnCode <> #old.pnCode[#pStn].me THEN

                   REGION "SET FLAG"
                       #ret := TRUE;
                   END_REGION

               END_IF;
           END_REGION

           REGION "SAVE FLAG"
               #stns.stn[#pStn].wipCmpts.flags.newPN := #ret;
           END_REGION

           REGION "CHANGE DETECTION"
               #old.pnCode[#pStn].me := #stns.stn[#pStn].wipCmpts.pnCode;
           END_REGION

       END_FOR;
   END_REGION
END_FUNCTION_BLOCK

FUNCTION_BLOCK "Flag: State Transition"   // FB4, SCL
{ S7_Optimized_Access := 'TRUE' }
VERSION : 0.1
   VAR_IN_OUT
      stns : "Station: All Stations";
   END_VAR
   VAR
      old : Struct
         stn : Array[0.."stnCount"] of Struct
            orderState : Array[0.."btnCount"] of Int;
         END_STRUCT;
      END_STRUCT;
   END_VAR
   VAR_TEMP
      pStn : Int;
      pBtn : Int;
      ret : Bool;
   END_VAR
BEGIN
   REGION "FOR EACH STATION"
       FOR #pStn := 0 TO "stnCount" DO

           REGION "IGNORE WIP LOAD CYCLE"
               IF NOT #stns.stn[#pStn].flags.wipSwapped THEN

                   REGION "FOR EACH BUTTON"
                       FOR #pBtn := 0 TO "btnCount" DO

                           REGION "RESET RETURN"
                               #ret := FALSE;
                           END_REGION

                           REGION "ON CHANGE IN STATE"
                               IF #stns.stn[#pStn].wipCmpts.orderState[#pBtn] <> #old.stn[#pStn].orderState[#pBtn] THEN

                                   REGION "SET STATE TRANSITION FLAG"
                                       #ret := true;
                                   END_REGION

                               END_IF;
                           END_REGION

                           REGION "SAVE FLAG"
                               #stns.stn[#pStn].flags.stateTransition[#pBtn] := #ret;
                           END_REGION

                       END_FOR;
                   END_REGION

               END_IF;
           END_REGION

           REGION "CHANGE DETECTION"
               #old.stn[#pStn].orderState := #stns.stn[#pStn].wipCmpts.orderState;
           END_REGION

       END_FOR;
   END_REGION
END_FUNCTION_BLOCK

FUNCTION_BLOCK "Flag"   // FB5, SCL
{ S7_Optimized_Access := 'TRUE' }
VERSION : 0.1
   VAR_INPUT
      pnLib : "Recipe: PN Text Library";
   END_VAR
   VAR_IN_OUT
      stns : "Station: All Stations";
      savedStns : "Recipe: HMI Stations Saved Wips";
   END_VAR
   VAR
      "inst New PN Code" : "Flag: New PN Code";
      "inst Flag: State Transition" : "Flag: State Transition";
      "inst Flag: Wip Deselect" : "Flag: Wip Deselect";
      "inst Flag: Wip Swapped" : "Flag: Wip Swapped";
   END_VAR
BEGIN
   REGION "NEW PART NUMBER ASSIGNED"
       #"inst New PN Code"(#stns);
   END_REGION

   REGION "PART NUMBER VALIDATION"
       "Flag: PN Good"(pnLib := #pnLib,
                       stns := #stns);
   END_REGION

   REGION "WIP SWAPPED"
       #"inst Flag: Wip Swapped"(#stns);
   END_REGION

   REGION "STATE TRANSITIONS"
       #"inst Flag: State Transition"(#stns);
   END_REGION

   REGION "WIP DESELECTION"
       #"inst Flag: Wip Deselect"(#savedStns);
   END_REGION
END_FUNCTION_BLOCK

FUNCTION_BLOCK "Flag: Wip Swapped"   // FB10, SCL
{ S7_Optimized_Access := 'TRUE' }
VERSION : 0.1
   VAR_IN_OUT
      stns : "Station: All Stations";
   END_VAR
   VAR
      old : Struct
         wipIndex : Array[0.."stnCount"] of DInt;
      END_STRUCT;
   END_VAR
   VAR_TEMP
      pStn : Int;
      ret : Bool;
   END_VAR
BEGIN
   REGION "FOR EACH STATION"
       FOR #pStn := 0 TO "stnCount" DO

           REGION "ON WIP CHANGE"
               IF #stns.stn[#pStn].wipData.index <> #old.wipIndex[#pStn] THEN

                   REGION "SET FLAG"
                       #ret := TRUE;
                   END_REGION

                   REGION "SAVE FLAG"
                       #stns.stn[#pStn].wipCmpts.flags.newPN := #ret;
                   END_REGION

               END_IF;
           END_REGION

           REGION "CHANGE DETECTION"
               #old.wipIndex[#pStn] := #stns.stn[#pStn].wipData.index;
           END_REGION

       END_FOR;
   END_REGION
END_FUNCTION_BLOCK

FUNCTION_BLOCK "Flag: Wip Deselect: Flag Pulse"   // FB17, SCL
{ S7_Optimized_Access := 'TRUE' }
VERSION : 0.1
   VAR_INPUT
      remaining : Real;
      reset : Bool;
   END_VAR
   VAR_IN_OUT
      flag : Bool;
   END_VAR
   VAR RETAIN
      hasBeenFlipped : Bool;
   END_VAR
BEGIN
   #flag := FALSE;

   IF #reset THEN
       #hasBeenFlipped := FALSE;
       RETURN;
   END_IF;

   IF #remaining >= 0.0 THEN
       #hasBeenFlipped := FALSE;
       RETURN;
   END_IF;

   IF NOT #hasBeenFlipped THEN
       IF #remaining < 0.0 THEN
           #hasBeenFlipped := TRUE;
           #flag := TRUE;
       END_IF;
   END_IF;
END_FUNCTION_BLOCK

FUNCTION_BLOCK "Flag: Wip Deselect"   // FB18, SCL
{ S7_Optimized_Access := 'TRUE' }
VERSION : 0.1
   VAR_IN_OUT
      savedStns : "Recipe: HMI Stations Saved Wips";
   END_VAR
   VAR
      "inst Flag Pulses" : Array[0.."stnCount", 0.."wipCount"] of "Flag: Wip Deselect: Flag Pulse";
   END_VAR
   VAR_TEMP
      pStn : Int;
      pWip : Int;
   END_VAR
BEGIN
   REGION "FOR EACH STATION"
       FOR #pStn := 0 TO "hmi_station_count" DO

           REGION "FOR EACH WIP"
               FOR #pWip := 0 TO "wipCount" DO

                   REGION "FLAG PULSE"
                       #"inst Flag Pulses"[#pStn, #pWip](remaining := #savedStns.stn[#pStn].wip[#pWip].timers.wdsRemaining,
                                                         flag := #savedStns.stn[#pStn].wip[#pWip].flags.clearWipRequest);
                   END_REGION

               END_FOR;
           END_REGION

       END_FOR;
   END_REGION
END_FUNCTION_BLOCK

FUNCTION "Flag: PN Good" : Void   // FC13, SCL
{ S7_Optimized_Access := 'TRUE' }
VERSION : 0.1
   VAR_INPUT
      pnLib : "Recipe: PN Text Library";
   END_VAR
   VAR_IN_OUT
      stns : "Station: All Stations";
   END_VAR
   VAR_TEMP
      pStn : Int;
      pBtn : Int;
      pnGood : Bool;
   END_VAR
BEGIN
   REGION "FOR EACH STATION"
       FOR #pStn := 0 TO "stnCount" DO

           REGION "FOR EACH BUTTON"
               FOR #pBtn := 0 TO "btnCount" DO

                   REGION "ON NEW PN"
                       IF #stns.stn[#pStn].wipCmpts.flags.newPN THEN

                           REGION "VALIDATE PN"
                               #pnGood := "Validate PN"(pnCode := #stns.stn[#pStn].wipCmpts.pnCode[#pBtn],
                                                        pnLib := #pnLib);
                           END_REGION

                           REGION "SAVE TO FLAG"
                               #stns.stn[#pStn].wipCmpts.flags.pnGood[#pBtn] := #pnGood;
                           END_REGION

                       END_IF;
                   END_REGION

               END_FOR;
           END_REGION

       END_FOR;
   END_REGION
END_FUNCTION

// folder: From Excel

FUNCTION_BLOCK "From Excel"   // FB8, SCL
{ S7_Optimized_Access := 'TRUE' }
VERSION : 0.1
   VAR_INPUT
      codeLib : "From Excel: Data";
   END_VAR
   VAR_IN_OUT
      stns : "Station: All Stations";
      svdHMIStnWips : "Recipe: HMI Stations Saved Wips";
   END_VAR
   VAR
      codeToKP8Stn : Bool;
      codeToHMIStn : Bool;
      codeToSavedHMIStn : Bool;
      initializeHmiStations : Bool;
   END_VAR
BEGIN
   REGION "KP8 STATIONS"
       IF #codeToKP8Stn THEN
           "From Excel: PN Code to KP8 Stations"(codeLib := #codeLib,
                                                 stns := #stns);
       END_IF;
   END_REGION

   REGION "HMI STATIONS"
       IF #codeToHMIStn THEN
           "From Excel: PN Code to HMI Stations"(xlCodeLib := #codeLib,
                                                 stns := #stns);
       END_IF;
   END_REGION


   REGION "SAVED HMI STATION WIPS"
       IF #codeToSavedHMIStn THEN
           "From Excel: PN Code to HMI Station Saved Wips"(codeLib := #codeLib,
                                                           savedWipStns := #svdHMIStnWips);
           "From Excel: Wip Code to HMI Station Saved WIps"(xlCodeLib := #codeLib,
                                                            savedWipStns := #svdHMIStnWips);
       END_IF;
   END_REGION

   REGION "MANUALLY STARTUP ROUTINE"
       IF #initializeHmiStations THEN
           "HMI Station Initialization"();
       END_IF;
   END_REGION
END_FUNCTION_BLOCK

FUNCTION "From Excel: PN Code to KP8 Stations" : Void   // FC58, SCL
{ S7_Optimized_Access := 'TRUE' }
VERSION : 0.1
   VAR_INPUT
      codeLib : "From Excel: Data";
   END_VAR
   VAR_IN_OUT
      stns : "Station: All Stations";
   END_VAR
   VAR_TEMP
      pSrc : Int;
      pDest : Int;
   END_VAR
BEGIN
   REGION "KP8 STATIONS
       FOR #pSrc := 0 TO UDINT_TO_INT("Length"(#codeLib.kp8Stns) - 1) DO
           #pDest := #codeLib.kp8Stns[#pSrc].pStn;
           IF #pDest = -1 THEN
               EXIT;
           END_IF;
           #stns.stn[#pDest].wipCmpts.pnCode := #codeLib.kp8Stns[#pSrc].pnCode;
       END_FOR;
   END_REGION
END_FUNCTION
